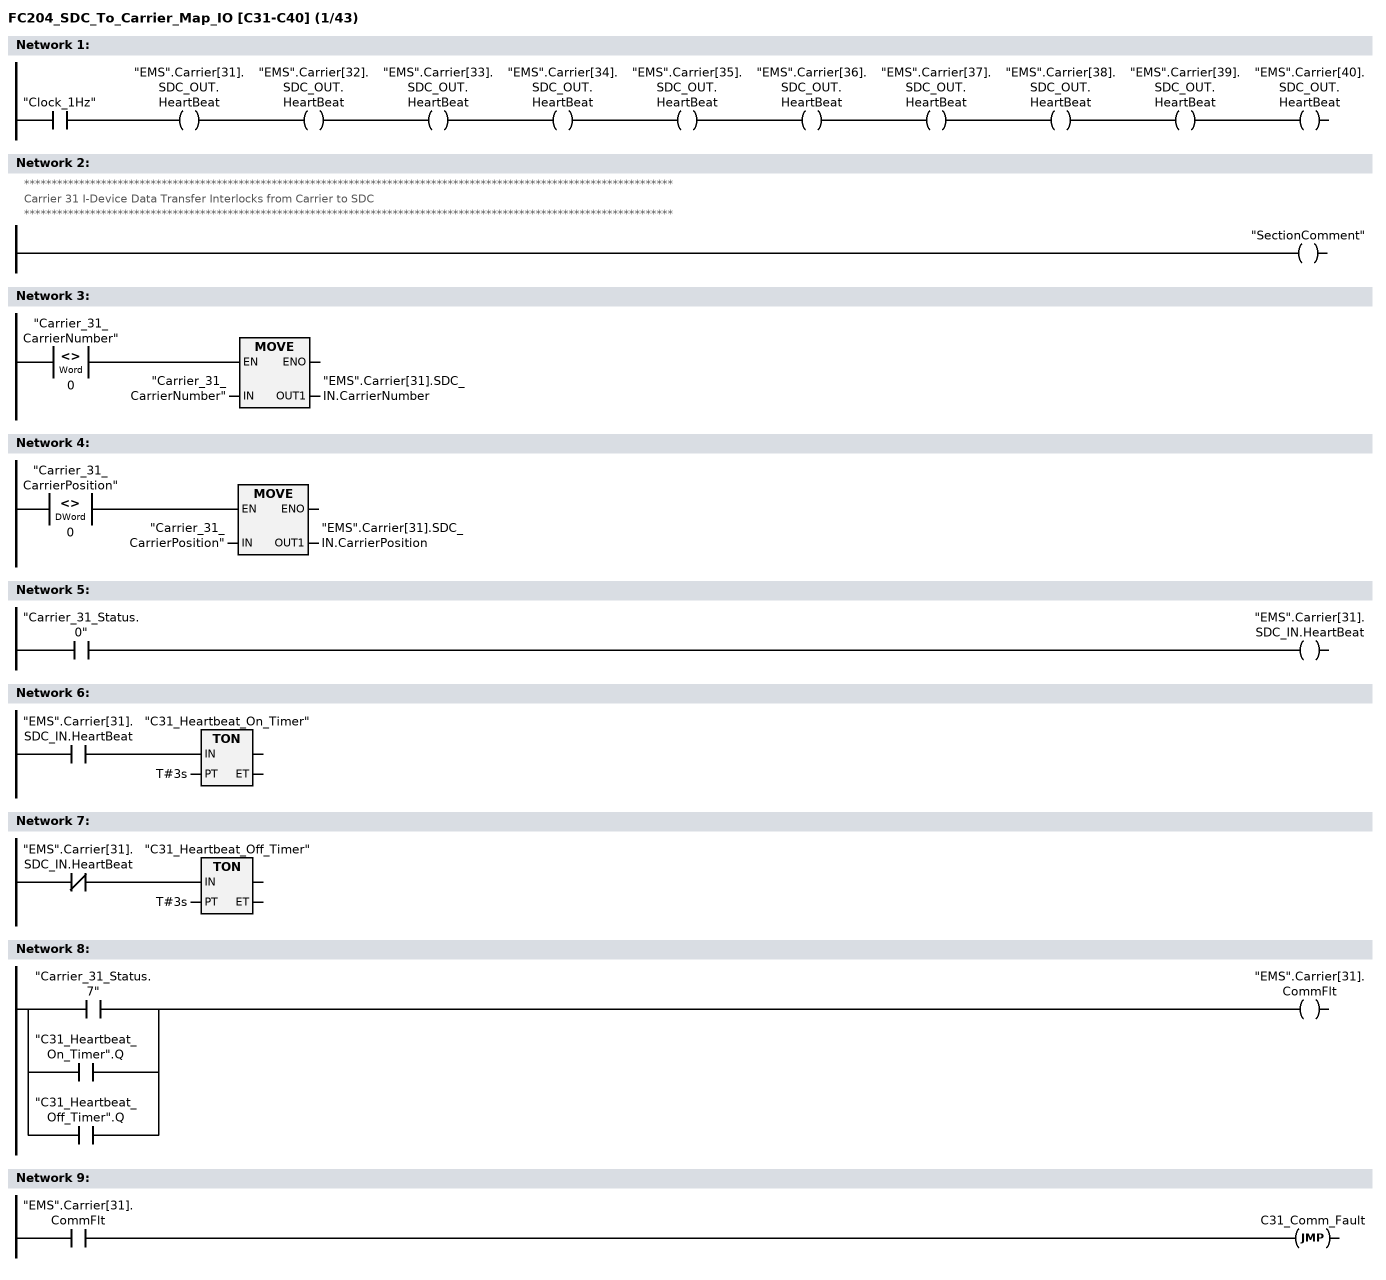
   RUNG wire#powerrail
      Contact( "Clock_1Hz" )
      Coil( "EMS".Carrier[31].SDC_OUT.HeartBeat )
      Coil( "EMS".Carrier[32].SDC_OUT.HeartBeat )
      Coil( "EMS".Carrier[33].SDC_OUT.HeartBeat )
      Coil( "EMS".Carrier[34].SDC_OUT.HeartBeat )
      Coil( "EMS".Carrier[35].SDC_OUT.HeartBeat )
      Coil( "EMS".Carrier[36].SDC_OUT.HeartBeat )
      Coil( "EMS".Carrier[37].SDC_OUT.HeartBeat )
      Coil( "EMS".Carrier[38].SDC_OUT.HeartBeat )
      Coil( "EMS".Carrier[39].SDC_OUT.HeartBeat )
      Coil( "EMS".Carrier[40].SDC_OUT.HeartBeat )
   END_RUNG
   // the same network as SCL:
   "EMS".Carrier[31].SDC_OUT.HeartBeat := "Clock_1Hz";
   "EMS".Carrier[32].SDC_OUT.HeartBeat := "Clock_1Hz";
   "EMS".Carrier[33].SDC_OUT.HeartBeat := "Clock_1Hz";
   "EMS".Carrier[34].SDC_OUT.HeartBeat := "Clock_1Hz";
   "EMS".Carrier[35].SDC_OUT.HeartBeat := "Clock_1Hz";
   "EMS".Carrier[36].SDC_OUT.HeartBeat := "Clock_1Hz";
   "EMS".Carrier[37].SDC_OUT.HeartBeat := "Clock_1Hz";
   "EMS".Carrier[38].SDC_OUT.HeartBeat := "Clock_1Hz";
   "EMS".Carrier[39].SDC_OUT.HeartBeat := "Clock_1Hz";
   "EMS".Carrier[40].SDC_OUT.HeartBeat := "Clock_1Hz";
END_REGION

REGION Network 2
   // **********************************************************************************************************************
   // 
   // Carrier 31 I-Device Data Transfer Interlocks from Carrier to SDC
   // 
   // **********************************************************************************************************************
   RUNG wire#powerrail
      Coil( "SectionComment" )
   END_RUNG
   // the same network as SCL:
   "SectionComment" := TRUE;
END_REGION

REGION Network 3
   RUNG wire#powerrail
      { S7_Templates := "SrcType := Word" } NE_Contact(in1 := "Carrier_31_CarrierNumber", in2 := 0)
      Move(in := "Carrier_31_CarrierNumber", out1 => "EMS".Carrier[31].SDC_IN.CarrierNumber)
   END_RUNG
   // the same network as SCL:
   IF "Carrier_31_CarrierNumber" <> 0 THEN
       "EMS".Carrier[31].SDC_IN.CarrierNumber := "Carrier_31_CarrierNumber";
   END_IF;
END_REGION

REGION Network 4
   RUNG wire#powerrail
      { S7_Templates := "SrcType := DWord" } NE_Contact(in1 := "Carrier_31_CarrierPosition", in2 := 0)
      Move(in := "Carrier_31_CarrierPosition", out1 => "EMS".Carrier[31].SDC_IN.CarrierPosition)
   END_RUNG
   // the same network as SCL:
   IF "Carrier_31_CarrierPosition" <> 0 THEN
       "EMS".Carrier[31].SDC_IN.CarrierPosition := "Carrier_31_CarrierPosition";
   END_IF;
END_REGION

REGION Network 5
   RUNG wire#powerrail
      Contact( "Carrier_31_Status.0" )
      Coil( "EMS".Carrier[31].SDC_IN.HeartBeat )
   END_RUNG
   // the same network as SCL:
   "EMS".Carrier[31].SDC_IN.HeartBeat := "Carrier_31_Status.0";
END_REGION

REGION Network 6
   "C31_Heartbeat_On_Timer".TON(IN := "EMS".Carrier[31].SDC_IN.HeartBeat, PT := T#3s);
END_REGION

REGION Network 7
   "C31_Heartbeat_Off_Timer".TON(IN := NOT "EMS".Carrier[31].SDC_IN.HeartBeat, PT := T#3s);
END_REGION

REGION Network 8
   RUNG wire#powerrail
      Contact( "Carrier_31_Status.7" )
      wire#w1
      Coil( "EMS".Carrier[31].CommFlt )
   END_RUNG
   RUNG wire#powerrail
      Contact( "C31_Heartbeat_On_Timer".Q )
   END_RUNG wire#w1
   RUNG wire#powerrail
      Contact( "C31_Heartbeat_Off_Timer".Q )
   END_RUNG wire#w1
   // the same network as SCL:
   "EMS".Carrier[31].CommFlt := "Carrier_31_Status.7" OR "C31_Heartbeat_On_Timer".Q OR "C31_Heartbeat_Off_Timer".Q;
END_REGION

REGION Network 9
   RUNG wire#powerrail
      Contact( "EMS".Carrier[31].CommFlt )
      JumpCoil( C31_Comm_Fault )
   END_RUNG
   // the same network as SCL:
   IF "EMS".Carrier[31].CommFlt THEN GOTO C31_Comm_Fault; END_IF;
END_REGION

REGION Network 10
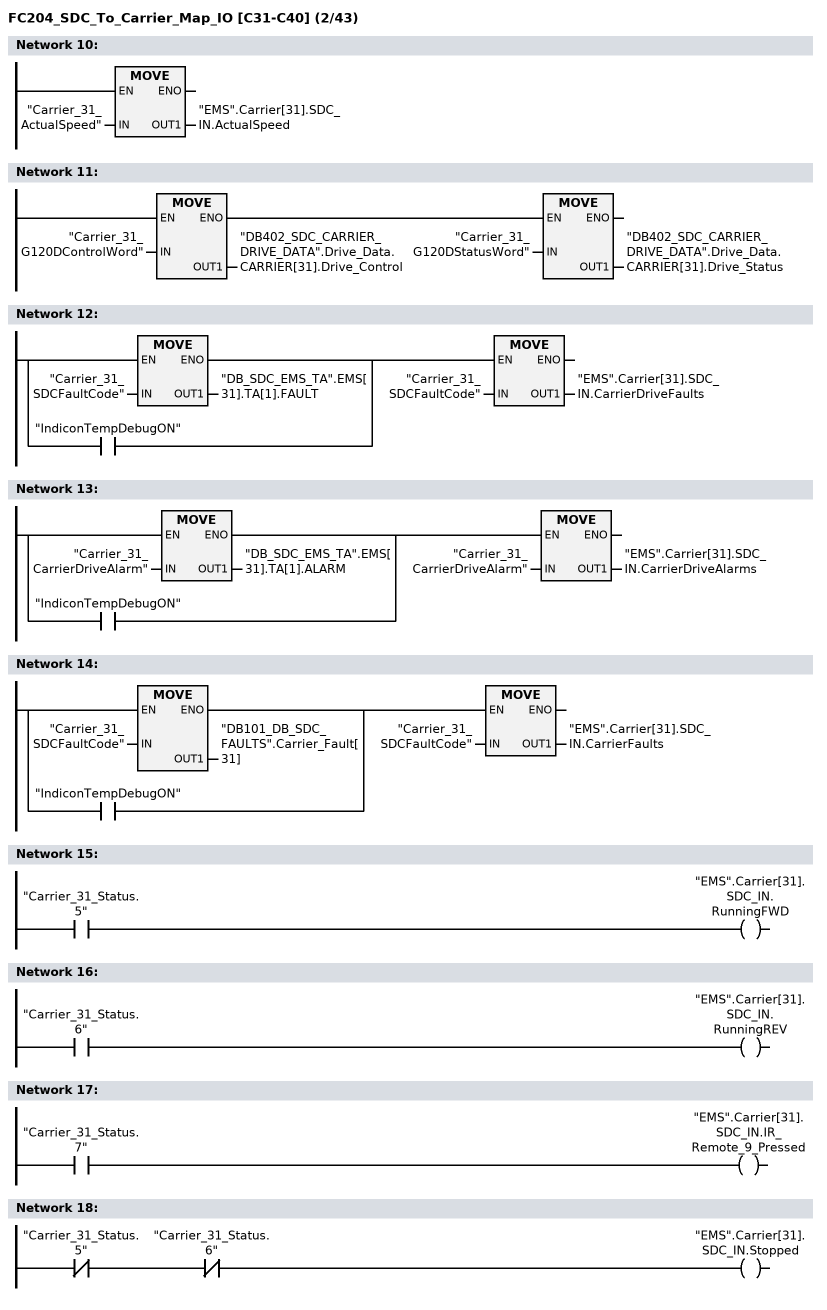
   RUNG wire#powerrail
      Move(in := "Carrier_31_ActualSpeed", out1 => "EMS".Carrier[31].SDC_IN.ActualSpeed)
   END_RUNG
   // the same network as SCL:
   "EMS".Carrier[31].SDC_IN.ActualSpeed := "Carrier_31_ActualSpeed";
END_REGION

REGION Network 11
   RUNG wire#powerrail
      Move(in := "Carrier_31_G120DControlWord", out1 => "DB402_SDC_CARRIER_DRIVE_DATA".Drive_Data.CARRIER[31].Drive_Control)
      Move(in := "Carrier_31_G120DStatusWord", out1 => "DB402_SDC_CARRIER_DRIVE_DATA".Drive_Data.CARRIER[31].Drive_Status)
   END_RUNG
   // the same network as SCL:
   "DB402_SDC_CARRIER_DRIVE_DATA".Drive_Data.CARRIER[31].Drive_Control := "Carrier_31_G120DControlWord";
   "DB402_SDC_CARRIER_DRIVE_DATA".Drive_Data.CARRIER[31].Drive_Status := "Carrier_31_G120DStatusWord";
END_REGION

REGION Network 12
   RUNG wire#powerrail
      Move(in := "Carrier_31_SDCFaultCode", out1 => "DB_SDC_EMS_TA".EMS[31].TA[1].FAULT)
      wire#w1
      Move(in := "Carrier_31_SDCFaultCode", out1 => "EMS".Carrier[31].SDC_IN.CarrierDriveFaults)
   END_RUNG
   RUNG wire#powerrail
      Contact( "IndiconTempDebugON" )
   END_RUNG wire#w1
   // the same network as SCL:
   "DB_SDC_EMS_TA".EMS[31].TA[1].FAULT := "Carrier_31_SDCFaultCode";
   IF TRUE OR "IndiconTempDebugON" THEN
       "EMS".Carrier[31].SDC_IN.CarrierDriveFaults := "Carrier_31_SDCFaultCode";
   END_IF;
END_REGION

REGION Network 13
   RUNG wire#powerrail
      Move(in := "Carrier_31_CarrierDriveAlarm", out1 => "DB_SDC_EMS_TA".EMS[31].TA[1].ALARM)
      wire#w1
      Move(in := "Carrier_31_CarrierDriveAlarm", out1 => "EMS".Carrier[31].SDC_IN.CarrierDriveAlarms)
   END_RUNG
   RUNG wire#powerrail
      Contact( "IndiconTempDebugON" )
   END_RUNG wire#w1
   // the same network as SCL:
   "DB_SDC_EMS_TA".EMS[31].TA[1].ALARM := "Carrier_31_CarrierDriveAlarm";
   IF TRUE OR "IndiconTempDebugON" THEN
       "EMS".Carrier[31].SDC_IN.CarrierDriveAlarms := "Carrier_31_CarrierDriveAlarm";
   END_IF;
END_REGION

REGION Network 14
   RUNG wire#powerrail
      Move(in := "Carrier_31_SDCFaultCode", out1 => "DB101_DB_SDC_FAULTS".Carrier_Fault[31])
      wire#w1
      Move(in := "Carrier_31_SDCFaultCode", out1 => "EMS".Carrier[31].SDC_IN.CarrierFaults)
   END_RUNG
   RUNG wire#powerrail
      Contact( "IndiconTempDebugON" )
   END_RUNG wire#w1
   // the same network as SCL:
   "DB101_DB_SDC_FAULTS".Carrier_Fault[31] := "Carrier_31_SDCFaultCode";
   IF TRUE OR "IndiconTempDebugON" THEN
       "EMS".Carrier[31].SDC_IN.CarrierFaults := "Carrier_31_SDCFaultCode";
   END_IF;
END_REGION

REGION Network 15
   RUNG wire#powerrail
      Contact( "Carrier_31_Status.5" )
      Coil( "EMS".Carrier[31].SDC_IN.RunningFWD )
   END_RUNG
   // the same network as SCL:
   "EMS".Carrier[31].SDC_IN.RunningFWD := "Carrier_31_Status.5";
END_REGION

REGION Network 16
   RUNG wire#powerrail
      Contact( "Carrier_31_Status.6" )
      Coil( "EMS".Carrier[31].SDC_IN.RunningREV )
   END_RUNG
   // the same network as SCL:
   "EMS".Carrier[31].SDC_IN.RunningREV := "Carrier_31_Status.6";
END_REGION

REGION Network 17
   RUNG wire#powerrail
      Contact( "Carrier_31_Status.7" )
      Coil( "EMS".Carrier[31].SDC_IN.IR_Remote_9_Pressed )
   END_RUNG
   // the same network as SCL:
   "EMS".Carrier[31].SDC_IN.IR_Remote_9_Pressed := "Carrier_31_Status.7";
END_REGION

REGION Network 18
   RUNG wire#powerrail
      I_Contact( "Carrier_31_Status.5" )
      I_Contact( "Carrier_31_Status.6" )
      Coil( "EMS".Carrier[31].SDC_IN.Stopped )
   END_RUNG
   // the same network as SCL:
   "EMS".Carrier[31].SDC_IN.Stopped := NOT "Carrier_31_Status.5" AND NOT "Carrier_31_Status.6";
END_REGION

REGION Network 19
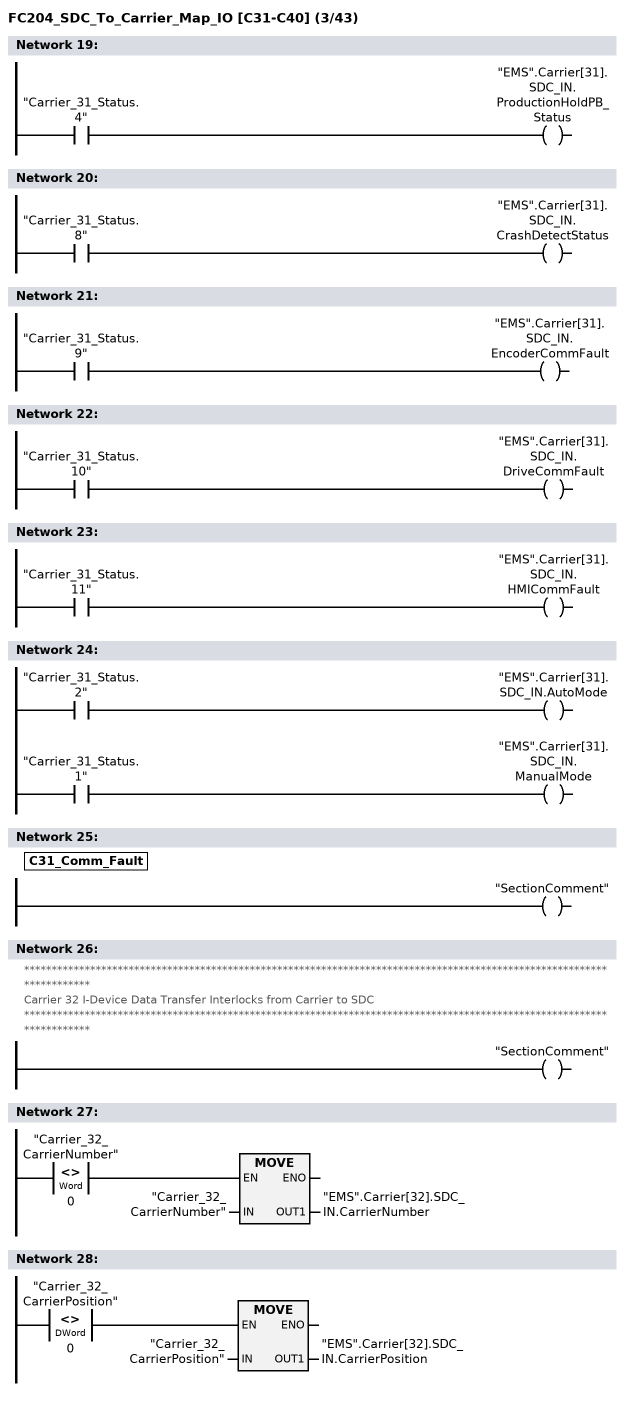
   RUNG wire#powerrail
      Contact( "Carrier_31_Status.4" )
      Coil( "EMS".Carrier[31].SDC_IN.ProductionHoldPB_Status )
   END_RUNG
   // the same network as SCL:
   "EMS".Carrier[31].SDC_IN.ProductionHoldPB_Status := "Carrier_31_Status.4";
END_REGION

REGION Network 20
   RUNG wire#powerrail
      Contact( "Carrier_31_Status.8" )
      Coil( "EMS".Carrier[31].SDC_IN.CrashDetectStatus )
   END_RUNG
   // the same network as SCL:
   "EMS".Carrier[31].SDC_IN.CrashDetectStatus := "Carrier_31_Status.8";
END_REGION

REGION Network 21
   RUNG wire#powerrail
      Contact( "Carrier_31_Status.9" )
      Coil( "EMS".Carrier[31].SDC_IN.EncoderCommFault )
   END_RUNG
   // the same network as SCL:
   "EMS".Carrier[31].SDC_IN.EncoderCommFault := "Carrier_31_Status.9";
END_REGION

REGION Network 22
   RUNG wire#powerrail
      Contact( "Carrier_31_Status.10" )
      Coil( "EMS".Carrier[31].SDC_IN.DriveCommFault )
   END_RUNG
   // the same network as SCL:
   "EMS".Carrier[31].SDC_IN.DriveCommFault := "Carrier_31_Status.10";
END_REGION

REGION Network 23
   RUNG wire#powerrail
      Contact( "Carrier_31_Status.11" )
      Coil( "EMS".Carrier[31].SDC_IN.HMICommFault )
   END_RUNG
   // the same network as SCL:
   "EMS".Carrier[31].SDC_IN.HMICommFault := "Carrier_31_Status.11";
END_REGION

REGION Network 24
   RUNG wire#powerrail
      Contact( "Carrier_31_Status.2" )
      Coil( "EMS".Carrier[31].SDC_IN.AutoMode )
   END_RUNG
   RUNG wire#powerrail
      Contact( "Carrier_31_Status.1" )
      Coil( "EMS".Carrier[31].SDC_IN.ManualMode )
   END_RUNG
   // the same network as SCL:
   "EMS".Carrier[31].SDC_IN.AutoMode := "Carrier_31_Status.2";
   "EMS".Carrier[31].SDC_IN.ManualMode := "Carrier_31_Status.1";
END_REGION

REGION Network 25
   Label( C31_Comm_Fault )
   RUNG wire#powerrail
      Coil( "SectionComment" )
   END_RUNG
   // the same network as SCL:
   C31_Comm_Fault:
   "SectionComment" := TRUE;
END_REGION

REGION Network 26
   // **********************************************************************************************************************
   // 
   // Carrier 32 I-Device Data Transfer Interlocks from Carrier to SDC
   // 
   // **********************************************************************************************************************
   RUNG wire#powerrail
      Coil( "SectionComment" )
   END_RUNG
   // the same network as SCL:
   "SectionComment" := TRUE;
END_REGION

REGION Network 27
   RUNG wire#powerrail
      { S7_Templates := "SrcType := Word" } NE_Contact(in1 := "Carrier_32_CarrierNumber", in2 := 0)
      Move(in := "Carrier_32_CarrierNumber", out1 => "EMS".Carrier[32].SDC_IN.CarrierNumber)
   END_RUNG
   // the same network as SCL:
   IF "Carrier_32_CarrierNumber" <> 0 THEN
       "EMS".Carrier[32].SDC_IN.CarrierNumber := "Carrier_32_CarrierNumber";
   END_IF;
END_REGION

REGION Network 28
   RUNG wire#powerrail
      { S7_Templates := "SrcType := DWord" } NE_Contact(in1 := "Carrier_32_CarrierPosition", in2 := 0)
      Move(in := "Carrier_32_CarrierPosition", out1 => "EMS".Carrier[32].SDC_IN.CarrierPosition)
   END_RUNG
   // the same network as SCL:
   IF "Carrier_32_CarrierPosition" <> 0 THEN
       "EMS".Carrier[32].SDC_IN.CarrierPosition := "Carrier_32_CarrierPosition";
   END_IF;
END_REGION

REGION Network 29
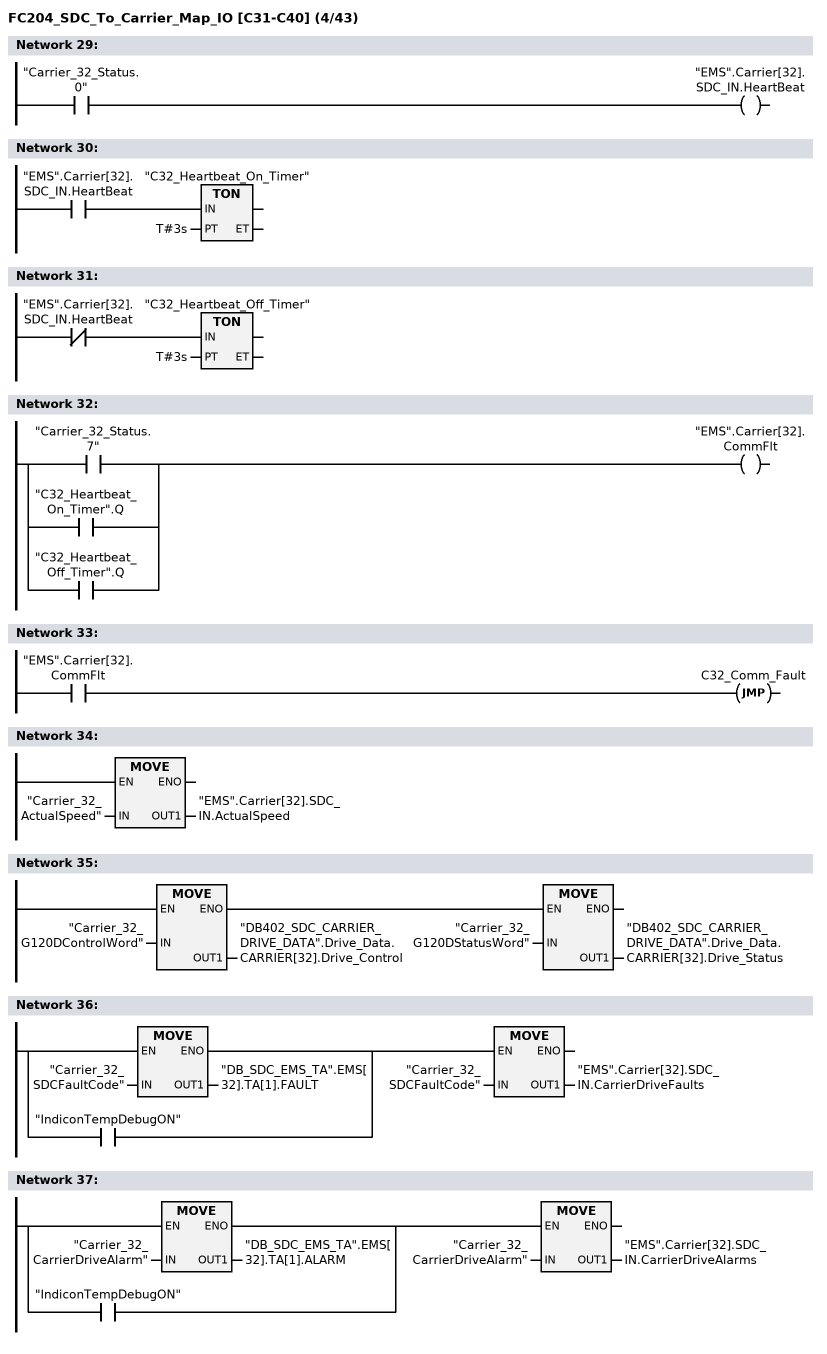
   RUNG wire#powerrail
      Contact( "Carrier_32_Status.0" )
      Coil( "EMS".Carrier[32].SDC_IN.HeartBeat )
   END_RUNG
   // the same network as SCL:
   "EMS".Carrier[32].SDC_IN.HeartBeat := "Carrier_32_Status.0";
END_REGION

REGION Network 30
   "C32_Heartbeat_On_Timer".TON(IN := "EMS".Carrier[32].SDC_IN.HeartBeat, PT := T#3s);
END_REGION

REGION Network 31
   "C32_Heartbeat_Off_Timer".TON(IN := NOT "EMS".Carrier[32].SDC_IN.HeartBeat, PT := T#3s);
END_REGION

REGION Network 32
   RUNG wire#powerrail
      Contact( "Carrier_32_Status.7" )
      wire#w1
      Coil( "EMS".Carrier[32].CommFlt )
   END_RUNG
   RUNG wire#powerrail
      Contact( "C32_Heartbeat_On_Timer".Q )
   END_RUNG wire#w1
   RUNG wire#powerrail
      Contact( "C32_Heartbeat_Off_Timer".Q )
   END_RUNG wire#w1
   // the same network as SCL:
   "EMS".Carrier[32].CommFlt := "Carrier_32_Status.7" OR "C32_Heartbeat_On_Timer".Q OR "C32_Heartbeat_Off_Timer".Q;
END_REGION

REGION Network 33
   RUNG wire#powerrail
      Contact( "EMS".Carrier[32].CommFlt )
      JumpCoil( C32_Comm_Fault )
   END_RUNG
   // the same network as SCL:
   IF "EMS".Carrier[32].CommFlt THEN GOTO C32_Comm_Fault; END_IF;
END_REGION

REGION Network 34
   RUNG wire#powerrail
      Move(in := "Carrier_32_ActualSpeed", out1 => "EMS".Carrier[32].SDC_IN.ActualSpeed)
   END_RUNG
   // the same network as SCL:
   "EMS".Carrier[32].SDC_IN.ActualSpeed := "Carrier_32_ActualSpeed";
END_REGION

REGION Network 35
   RUNG wire#powerrail
      Move(in := "Carrier_32_G120DControlWord", out1 => "DB402_SDC_CARRIER_DRIVE_DATA".Drive_Data.CARRIER[32].Drive_Control)
      Move(in := "Carrier_32_G120DStatusWord", out1 => "DB402_SDC_CARRIER_DRIVE_DATA".Drive_Data.CARRIER[32].Drive_Status)
   END_RUNG
   // the same network as SCL:
   "DB402_SDC_CARRIER_DRIVE_DATA".Drive_Data.CARRIER[32].Drive_Control := "Carrier_32_G120DControlWord";
   "DB402_SDC_CARRIER_DRIVE_DATA".Drive_Data.CARRIER[32].Drive_Status := "Carrier_32_G120DStatusWord";
END_REGION

REGION Network 36
   RUNG wire#powerrail
      Move(in := "Carrier_32_SDCFaultCode", out1 => "DB_SDC_EMS_TA".EMS[32].TA[1].FAULT)
      wire#w1
      Move(in := "Carrier_32_SDCFaultCode", out1 => "EMS".Carrier[32].SDC_IN.CarrierDriveFaults)
   END_RUNG
   RUNG wire#powerrail
      Contact( "IndiconTempDebugON" )
   END_RUNG wire#w1
   // the same network as SCL:
   "DB_SDC_EMS_TA".EMS[32].TA[1].FAULT := "Carrier_32_SDCFaultCode";
   IF TRUE OR "IndiconTempDebugON" THEN
       "EMS".Carrier[32].SDC_IN.CarrierDriveFaults := "Carrier_32_SDCFaultCode";
   END_IF;
END_REGION

REGION Network 37
   RUNG wire#powerrail
      Move(in := "Carrier_32_CarrierDriveAlarm", out1 => "DB_SDC_EMS_TA".EMS[32].TA[1].ALARM)
      wire#w1
      Move(in := "Carrier_32_CarrierDriveAlarm", out1 => "EMS".Carrier[32].SDC_IN.CarrierDriveAlarms)
   END_RUNG
   RUNG wire#powerrail
      Contact( "IndiconTempDebugON" )
   END_RUNG wire#w1
   // the same network as SCL:
   "DB_SDC_EMS_TA".EMS[32].TA[1].ALARM := "Carrier_32_CarrierDriveAlarm";
   IF TRUE OR "IndiconTempDebugON" THEN
       "EMS".Carrier[32].SDC_IN.CarrierDriveAlarms := "Carrier_32_CarrierDriveAlarm";
   END_IF;
END_REGION

REGION Network 38
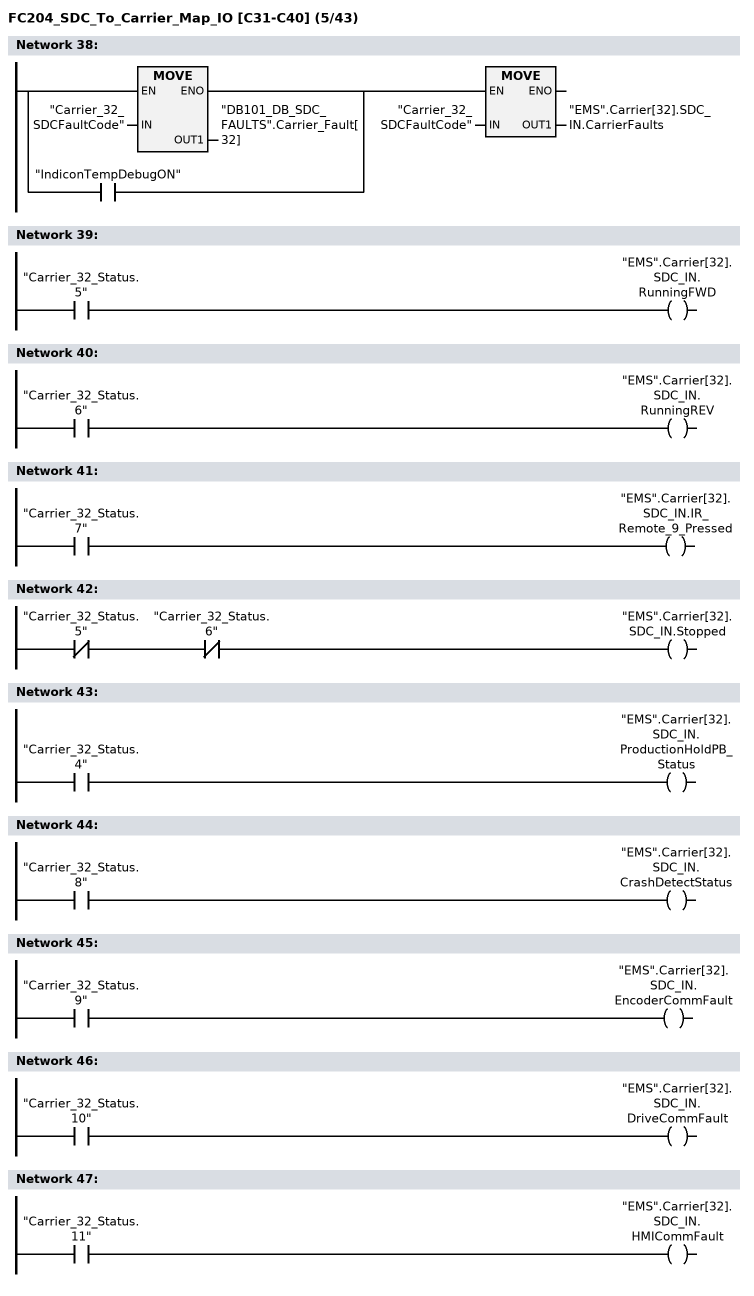
   RUNG wire#powerrail
      Move(in := "Carrier_32_SDCFaultCode", out1 => "DB101_DB_SDC_FAULTS".Carrier_Fault[32])
      wire#w1
      Move(in := "Carrier_32_SDCFaultCode", out1 => "EMS".Carrier[32].SDC_IN.CarrierFaults)
   END_RUNG
   RUNG wire#powerrail
      Contact( "IndiconTempDebugON" )
   END_RUNG wire#w1
   // the same network as SCL:
   "DB101_DB_SDC_FAULTS".Carrier_Fault[32] := "Carrier_32_SDCFaultCode";
   IF TRUE OR "IndiconTempDebugON" THEN
       "EMS".Carrier[32].SDC_IN.CarrierFaults := "Carrier_32_SDCFaultCode";
   END_IF;
END_REGION

REGION Network 39
   RUNG wire#powerrail
      Contact( "Carrier_32_Status.5" )
      Coil( "EMS".Carrier[32].SDC_IN.RunningFWD )
   END_RUNG
   // the same network as SCL:
   "EMS".Carrier[32].SDC_IN.RunningFWD := "Carrier_32_Status.5";
END_REGION

REGION Network 40
   RUNG wire#powerrail
      Contact( "Carrier_32_Status.6" )
      Coil( "EMS".Carrier[32].SDC_IN.RunningREV )
   END_RUNG
   // the same network as SCL:
   "EMS".Carrier[32].SDC_IN.RunningREV := "Carrier_32_Status.6";
END_REGION

REGION Network 41
   RUNG wire#powerrail
      Contact( "Carrier_32_Status.7" )
      Coil( "EMS".Carrier[32].SDC_IN.IR_Remote_9_Pressed )
   END_RUNG
   // the same network as SCL:
   "EMS".Carrier[32].SDC_IN.IR_Remote_9_Pressed := "Carrier_32_Status.7";
END_REGION

REGION Network 42
   RUNG wire#powerrail
      I_Contact( "Carrier_32_Status.5" )
      I_Contact( "Carrier_32_Status.6" )
      Coil( "EMS".Carrier[32].SDC_IN.Stopped )
   END_RUNG
   // the same network as SCL:
   "EMS".Carrier[32].SDC_IN.Stopped := NOT "Carrier_32_Status.5" AND NOT "Carrier_32_Status.6";
END_REGION

REGION Network 43
   RUNG wire#powerrail
      Contact( "Carrier_32_Status.4" )
      Coil( "EMS".Carrier[32].SDC_IN.ProductionHoldPB_Status )
   END_RUNG
   // the same network as SCL:
   "EMS".Carrier[32].SDC_IN.ProductionHoldPB_Status := "Carrier_32_Status.4";
END_REGION

REGION Network 44
   RUNG wire#powerrail
      Contact( "Carrier_32_Status.8" )
      Coil( "EMS".Carrier[32].SDC_IN.CrashDetectStatus )
   END_RUNG
   // the same network as SCL:
   "EMS".Carrier[32].SDC_IN.CrashDetectStatus := "Carrier_32_Status.8";
END_REGION

REGION Network 45
   RUNG wire#powerrail
      Contact( "Carrier_32_Status.9" )
      Coil( "EMS".Carrier[32].SDC_IN.EncoderCommFault )
   END_RUNG
   // the same network as SCL:
   "EMS".Carrier[32].SDC_IN.EncoderCommFault := "Carrier_32_Status.9";
END_REGION

REGION Network 46
   RUNG wire#powerrail
      Contact( "Carrier_32_Status.10" )
      Coil( "EMS".Carrier[32].SDC_IN.DriveCommFault )
   END_RUNG
   // the same network as SCL:
   "EMS".Carrier[32].SDC_IN.DriveCommFault := "Carrier_32_Status.10";
END_REGION

REGION Network 47
   RUNG wire#powerrail
      Contact( "Carrier_32_Status.11" )
      Coil( "EMS".Carrier[32].SDC_IN.HMICommFault )
   END_RUNG
   // the same network as SCL:
   "EMS".Carrier[32].SDC_IN.HMICommFault := "Carrier_32_Status.11";
END_REGION

REGION Network 48
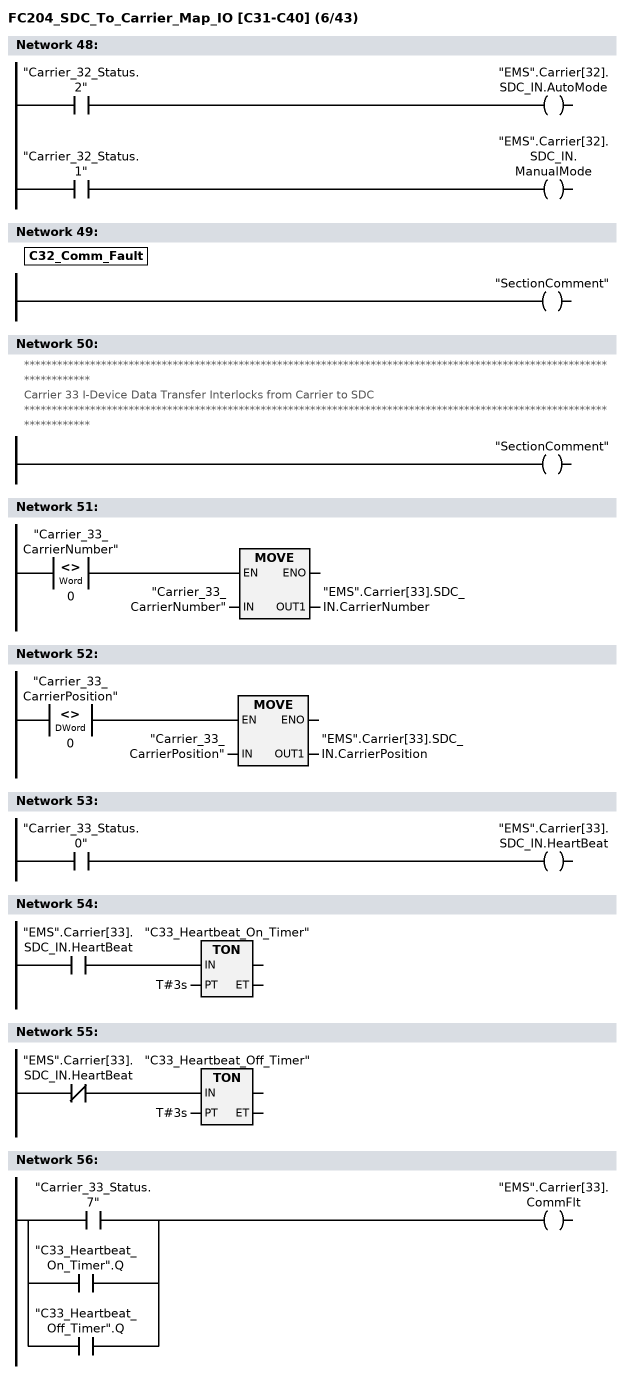
   RUNG wire#powerrail
      Contact( "Carrier_32_Status.2" )
      Coil( "EMS".Carrier[32].SDC_IN.AutoMode )
   END_RUNG
   RUNG wire#powerrail
      Contact( "Carrier_32_Status.1" )
      Coil( "EMS".Carrier[32].SDC_IN.ManualMode )
   END_RUNG
   // the same network as SCL:
   "EMS".Carrier[32].SDC_IN.AutoMode := "Carrier_32_Status.2";
   "EMS".Carrier[32].SDC_IN.ManualMode := "Carrier_32_Status.1";
END_REGION

REGION Network 49
   Label( C32_Comm_Fault )
   RUNG wire#powerrail
      Coil( "SectionComment" )
   END_RUNG
   // the same network as SCL:
   C32_Comm_Fault:
   "SectionComment" := TRUE;
END_REGION

REGION Network 50
   // **********************************************************************************************************************
   // 
   // Carrier 33 I-Device Data Transfer Interlocks from Carrier to SDC
   // 
   // **********************************************************************************************************************
   RUNG wire#powerrail
      Coil( "SectionComment" )
   END_RUNG
   // the same network as SCL:
   "SectionComment" := TRUE;
END_REGION

REGION Network 51
   RUNG wire#powerrail
      { S7_Templates := "SrcType := Word" } NE_Contact(in1 := "Carrier_33_CarrierNumber", in2 := 0)
      Move(in := "Carrier_33_CarrierNumber", out1 => "EMS".Carrier[33].SDC_IN.CarrierNumber)
   END_RUNG
   // the same network as SCL:
   IF "Carrier_33_CarrierNumber" <> 0 THEN
       "EMS".Carrier[33].SDC_IN.CarrierNumber := "Carrier_33_CarrierNumber";
   END_IF;
END_REGION

REGION Network 52
   RUNG wire#powerrail
      { S7_Templates := "SrcType := DWord" } NE_Contact(in1 := "Carrier_33_CarrierPosition", in2 := 0)
      Move(in := "Carrier_33_CarrierPosition", out1 => "EMS".Carrier[33].SDC_IN.CarrierPosition)
   END_RUNG
   // the same network as SCL:
   IF "Carrier_33_CarrierPosition" <> 0 THEN
       "EMS".Carrier[33].SDC_IN.CarrierPosition := "Carrier_33_CarrierPosition";
   END_IF;
END_REGION

REGION Network 53
   RUNG wire#powerrail
      Contact( "Carrier_33_Status.0" )
      Coil( "EMS".Carrier[33].SDC_IN.HeartBeat )
   END_RUNG
   // the same network as SCL:
   "EMS".Carrier[33].SDC_IN.HeartBeat := "Carrier_33_Status.0";
END_REGION

REGION Network 54
   "C33_Heartbeat_On_Timer".TON(IN := "EMS".Carrier[33].SDC_IN.HeartBeat, PT := T#3s);
END_REGION

REGION Network 55
   "C33_Heartbeat_Off_Timer".TON(IN := NOT "EMS".Carrier[33].SDC_IN.HeartBeat, PT := T#3s);
END_REGION

REGION Network 56
   RUNG wire#powerrail
      Contact( "Carrier_33_Status.7" )
      wire#w1
      Coil( "EMS".Carrier[33].CommFlt )
   END_RUNG
   RUNG wire#powerrail
      Contact( "C33_Heartbeat_On_Timer".Q )
   END_RUNG wire#w1
   RUNG wire#powerrail
      Contact( "C33_Heartbeat_Off_Timer".Q )
   END_RUNG wire#w1
   // the same network as SCL:
   "EMS".Carrier[33].CommFlt := "Carrier_33_Status.7" OR "C33_Heartbeat_On_Timer".Q OR "C33_Heartbeat_Off_Timer".Q;
END_REGION

REGION Network 57
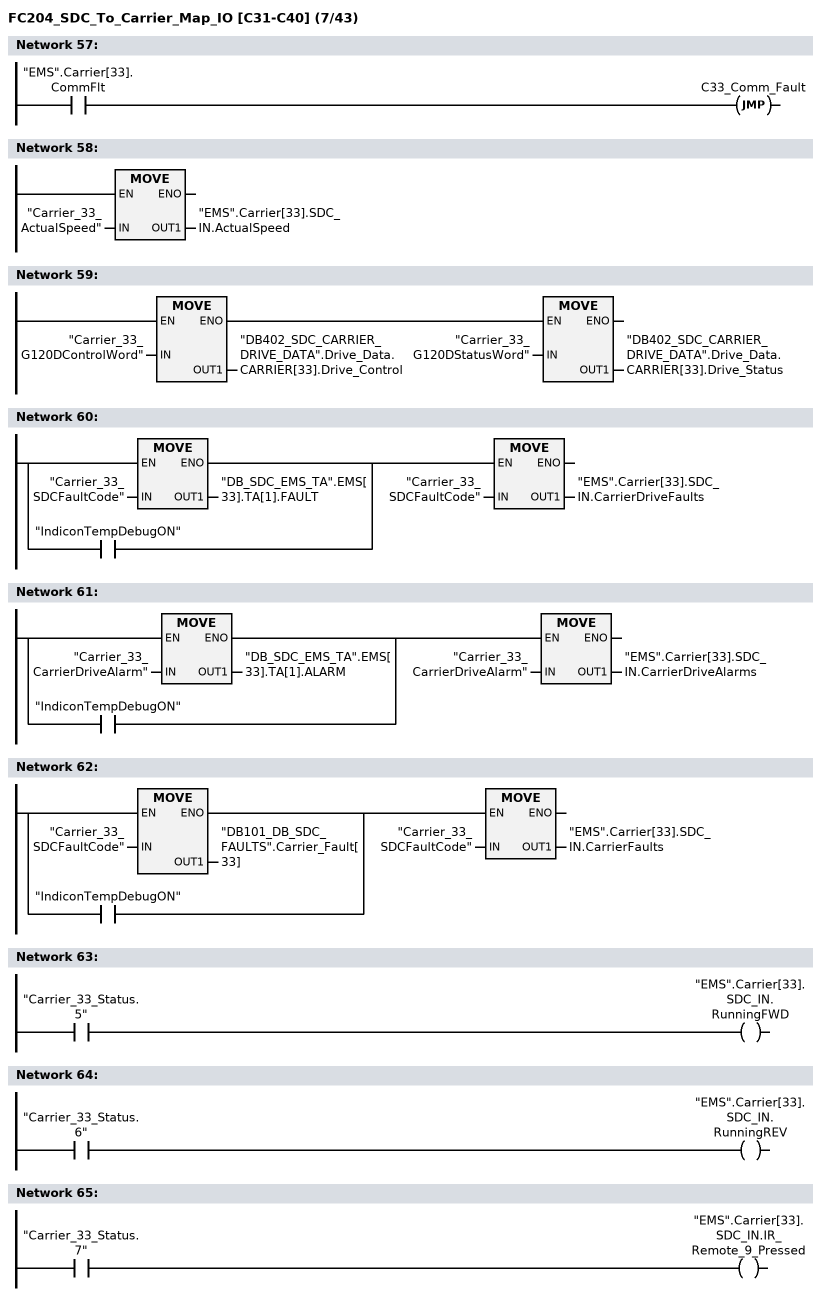
   RUNG wire#powerrail
      Contact( "EMS".Carrier[33].CommFlt )
      JumpCoil( C33_Comm_Fault )
   END_RUNG
   // the same network as SCL:
   IF "EMS".Carrier[33].CommFlt THEN GOTO C33_Comm_Fault; END_IF;
END_REGION

REGION Network 58
   RUNG wire#powerrail
      Move(in := "Carrier_33_ActualSpeed", out1 => "EMS".Carrier[33].SDC_IN.ActualSpeed)
   END_RUNG
   // the same network as SCL:
   "EMS".Carrier[33].SDC_IN.ActualSpeed := "Carrier_33_ActualSpeed";
END_REGION

REGION Network 59
   RUNG wire#powerrail
      Move(in := "Carrier_33_G120DControlWord", out1 => "DB402_SDC_CARRIER_DRIVE_DATA".Drive_Data.CARRIER[33].Drive_Control)
      Move(in := "Carrier_33_G120DStatusWord", out1 => "DB402_SDC_CARRIER_DRIVE_DATA".Drive_Data.CARRIER[33].Drive_Status)
   END_RUNG
   // the same network as SCL:
   "DB402_SDC_CARRIER_DRIVE_DATA".Drive_Data.CARRIER[33].Drive_Control := "Carrier_33_G120DControlWord";
   "DB402_SDC_CARRIER_DRIVE_DATA".Drive_Data.CARRIER[33].Drive_Status := "Carrier_33_G120DStatusWord";
END_REGION

REGION Network 60
   RUNG wire#powerrail
      Move(in := "Carrier_33_SDCFaultCode", out1 => "DB_SDC_EMS_TA".EMS[33].TA[1].FAULT)
      wire#w1
      Move(in := "Carrier_33_SDCFaultCode", out1 => "EMS".Carrier[33].SDC_IN.CarrierDriveFaults)
   END_RUNG
   RUNG wire#powerrail
      Contact( "IndiconTempDebugON" )
   END_RUNG wire#w1
   // the same network as SCL:
   "DB_SDC_EMS_TA".EMS[33].TA[1].FAULT := "Carrier_33_SDCFaultCode";
   IF TRUE OR "IndiconTempDebugON" THEN
       "EMS".Carrier[33].SDC_IN.CarrierDriveFaults := "Carrier_33_SDCFaultCode";
   END_IF;
END_REGION

REGION Network 61
   RUNG wire#powerrail
      Move(in := "Carrier_33_CarrierDriveAlarm", out1 => "DB_SDC_EMS_TA".EMS[33].TA[1].ALARM)
      wire#w1
      Move(in := "Carrier_33_CarrierDriveAlarm", out1 => "EMS".Carrier[33].SDC_IN.CarrierDriveAlarms)
   END_RUNG
   RUNG wire#powerrail
      Contact( "IndiconTempDebugON" )
   END_RUNG wire#w1
   // the same network as SCL:
   "DB_SDC_EMS_TA".EMS[33].TA[1].ALARM := "Carrier_33_CarrierDriveAlarm";
   IF TRUE OR "IndiconTempDebugON" THEN
       "EMS".Carrier[33].SDC_IN.CarrierDriveAlarms := "Carrier_33_CarrierDriveAlarm";
   END_IF;
END_REGION

REGION Network 62
   RUNG wire#powerrail
      Move(in := "Carrier_33_SDCFaultCode", out1 => "DB101_DB_SDC_FAULTS".Carrier_Fault[33])
      wire#w1
      Move(in := "Carrier_33_SDCFaultCode", out1 => "EMS".Carrier[33].SDC_IN.CarrierFaults)
   END_RUNG
   RUNG wire#powerrail
      Contact( "IndiconTempDebugON" )
   END_RUNG wire#w1
   // the same network as SCL:
   "DB101_DB_SDC_FAULTS".Carrier_Fault[33] := "Carrier_33_SDCFaultCode";
   IF TRUE OR "IndiconTempDebugON" THEN
       "EMS".Carrier[33].SDC_IN.CarrierFaults := "Carrier_33_SDCFaultCode";
   END_IF;
END_REGION

REGION Network 63
   RUNG wire#powerrail
      Contact( "Carrier_33_Status.5" )
      Coil( "EMS".Carrier[33].SDC_IN.RunningFWD )
   END_RUNG
   // the same network as SCL:
   "EMS".Carrier[33].SDC_IN.RunningFWD := "Carrier_33_Status.5";
END_REGION

REGION Network 64
   RUNG wire#powerrail
      Contact( "Carrier_33_Status.6" )
      Coil( "EMS".Carrier[33].SDC_IN.RunningREV )
   END_RUNG
   // the same network as SCL:
   "EMS".Carrier[33].SDC_IN.RunningREV := "Carrier_33_Status.6";
END_REGION

REGION Network 65
   RUNG wire#powerrail
      Contact( "Carrier_33_Status.7" )
      Coil( "EMS".Carrier[33].SDC_IN.IR_Remote_9_Pressed )
   END_RUNG
   // the same network as SCL:
   "EMS".Carrier[33].SDC_IN.IR_Remote_9_Pressed := "Carrier_33_Status.7";
END_REGION

REGION Network 66